VERSION : 0.1
// Die Funktion wird in einer Sprungleiste mit folgenden Schritten bearbeitet:
// 0: Warten, bis RT gedreht hat (nur danach ist Kettenentlastung notwendig)
// 1: Warten, bis BA Hand und keine Bewegung angefordert
// 2: Wartezeit vor Entlastung der Kette
//    -> Schritt 3, falls Wartezeit abgelaufen
//    -> Schritt 1, falls Automatik erneut angewählt oder Rundtisch dreht
// 3: Entlastung der Kette mit Zeitüberwachung
//    -> Schritt 1, falls während der Entlastung Bewegung angefordert wird
//    -> Schritt 0, falls während der Entlastung Automatik angewählt wird
// 4: Spannen der Kette mit Zeitüberwachung
   VAR_INPUT
      IN_P_Kette : Bool;   // Eingang von Druckschalter des Kettenspanners
      IN_Timer_Stg_Kette : Timer;   // Timer für die Störungsbildung der Spannung der Laufketten
      IN_Timer_Kettenspanner : Timer;   // Timer für den allgemeinen Ablauf des Kettenspanners
      IN_DW_Wartezeit : S5Time;   // Zeitwert für die Wartezeit nach Rundtisch im Handbetrieb
      IN_DW_Entlastungszeit : S5Time;   // Zeitwert für die Entlastungszeit der Kette
      IN_RT_dreht : Bool;   // Signal das sich der Rundtisch in Bewegung befindet
      IN_Steuerspannung : Bool;   // Signal Steuerspannung Eingeschaltet und Not- Aus entriegelt
      IN_Automatik_Stop_ok : Bool;   // Eingang das die Sicherheitseinrichtungen quittiert sind
      IN_Hydraulik_ok : Bool;   // Signal bei hydraulischen Kettenspannern das die Hydraulik bereit ist
      IN_Kettenspannung_noetig : Bool;   // Signal von extern das keine Kettenspannung nötig ist
      IN_Betriebsart_Automatik : Bool;   // Die Anlage befindet sich im Automatik- Betrieb
      IN_Start_Anlagenbetrieb : Bool;   // Die Anlage befindet sich in der Vorbereitung zum Produktionsbetrieb
      IN_Anlagenbetrieb : Bool;   // Die Anlage befindet sich im Produktionsbetrieb
      IN_Reset_fault_Fkt : Bool;   // Signal zum quittieren der Störungen innerhalb der einzelnen Funktionsbausteine
   END_VAR
   VAR_OUTPUT
      OUT_V_Entlastung : Bool;   // Ausgang für die Ansteuerung des Ketten- Entlastungs- Ventils
   END_VAR
   VAR_IN_OUT
      IO_Status : "UDT_RT_Kettenspanner";   // Speichern der Kettenentlastungs- Zustände für das Programm
   END_VAR
   VAR_TEMP
      Temp_IO_Status : "UDT_RT_Kettenspanner";   // Temporärer Kettenentlastungs- Status für die interne Bearbeitung des Bausteins
      ERROR_CODE : Int;   // Störungszustand der Systemfunktion "BLKMOV" Blockmove
      Anyzeiger : ANY;   // Zeiger zum Kopieren der Bereiche "IO_Status" und "Temp_IO_Status"
      Entlastung_starten : Bool;   // Zwischenmerker zum starten des Ablaufes der Kettenentspannung
   END_VAR
BEGIN

REGION Network 1: Gesicherte Daten einbinden
         LAR1;
         L;
         LAR2;
   //
         L     W#16#1002;  // Bytes
         T     W[AR1, P#0.0];
         L     2;  // Anzahl Bytes
         T     W[AR1, P#2.0];
         L     W[AR2, P#0.0];  // Baustein Nr.
         T     W[AR1, P#4.0];
         L     D[AR2, P#2.0];  // Datenanfang
         T     D[AR1, P#6.0];
   //
         CALL  BLKMOV
         ( SRCBLK  := #Anyzeiger,
           RET_VAL := #ERROR_CODE,
           DSTBLK  := #Temp_IO_Status
         );
   //
END_REGION

REGION Network 2: Stoerungen quittieren
         A     #IN_Reset_fault_Fkt;
         R     #Temp_IO_Status.STG_Entlastung;
         R     #Temp_IO_Status.STG_Druckaufbau;
END_REGION

REGION Network 3: Sprungleiste
         L     #Temp_IO_Status.Schrittnummer;
         JL    del;
         JU    dreh;  // 0: Warten, bis Rundtisch dreht
         JU    wrth;  // 1: Warten auf Betriebsart Hand + RT steht
         JU    wart;  // 2: Wartezeit vor Entlastung
         JU    entl;  // 3: Kettenentlastung
         JU    span;  // 4: Kette spannen
   del:  L     0;
         T     #Temp_IO_Status.Schrittnummer;
         CLR;
         =     #Temp_IO_Status.V_Entlastung;
         SP    #IN_Timer_Kettenspanner;
         SP    #IN_Timer_Stg_Kette;
         BEU;
END_REGION

REGION Network 4: 0: Warten, bis Rundtisch in Automatik gedreht hat
   dreh: ON    #IN_RT_dreht;
         ON    #IN_Anlagenbetrieb;
         JC    ende;
         L     1;
         T     #Temp_IO_Status.Schrittnummer;
         JU    ende;
END_REGION

REGION Network 5: 1: Warten, bis Automatik beendet und keine Bewegung läuft
   wrth: O     #IN_RT_dreht;
         O     #IN_Betriebsart_Automatik;
         JC    ende;
         L     2;
         T     #Temp_IO_Status.Schrittnummer;
         JU    ende;
END_REGION

REGION Network 6: 2: Wartezeit vor Kettenentlastung
   wart: SET;
         L     #IN_DW_Wartezeit;
         SD    #IN_Timer_Kettenspanner;
         L     1;
         O     #IN_RT_dreht;
         O     #IN_Start_Anlagenbetrieb;
         O     #IN_Anlagenbetrieb;
         JC    trnr;
         L     3;
         A     #IN_Timer_Kettenspanner;
         JC    trnr;
         JU    ende;
   trnr: T     #Temp_IO_Status.Schrittnummer;
         CLR;
         SP    #IN_Timer_Kettenspanner;
END_REGION

REGION Network 7: 3: Kettenentlastung
   entl: A     #IN_Steuerspannung;
         A     #IN_Automatik_Stop_ok;
         AN    #IN_RT_dreht;
         AN    #IN_Betriebsart_Automatik;
         AN    #IN_Kettenspannung_noetig;
         =     #Entlastung_starten;
         L     #IN_DW_Entlastungszeit;
         SP    #IN_Timer_Kettenspanner;
   //
         A     #Entlastung_starten;
         A     #IN_Timer_Kettenspanner;
         =     #Temp_IO_Status.V_Entlastung;
   //
         L     1;
         AN    #Entlastung_starten;
         JC    trn2;
         L     4;
         A     #Entlastung_starten;
         AN    #Temp_IO_Status.V_Entlastung;
         JC    trn2;
         JU    ende;
   trn2: T     #Temp_IO_Status.Schrittnummer;
         CLR;
         SP    #IN_Timer_Kettenspanner;
         JU    ende;
END_REGION

REGION Network 8: 4: Kette Spannen
   span: R     #Temp_IO_Status.V_Entlastung;
         L     0;
         T     #Temp_IO_Status.Schrittnummer;
END_REGION

REGION Network 9: Ende
   ende: A     #Temp_IO_Status.V_Entlastung;
         A     #IN_P_Kette;
         O;
         AN    #Temp_IO_Status.V_Entlastung;
         AN    #IN_P_Kette;
         A     #IN_Hydraulik_ok;
         L     S5T#10S;
         SD    #IN_Timer_Stg_Kette;
   //
         A     #IN_Timer_Stg_Kette;
         A     #Temp_IO_Status.V_Entlastung;
         S     #Temp_IO_Status.STG_Entlastung;
   //
         A     #IN_Timer_Stg_Kette;
         AN    #Temp_IO_Status.V_Entlastung;
         S     #Temp_IO_Status.STG_Druckaufbau;
   //
         AN    #Temp_IO_Status.V_Entlastung;
         A     #IN_P_Kette;
         =     #Temp_IO_Status.Kette_gespannt;
END_REGION

REGION Network 10: Ansteuerung des Entlanstungsventils
         A     #Temp_IO_Status.V_Entlastung;
         =     #OUT_V_Entlastung;
END_REGION

REGION Network 11: Daten sichern
         CALL  BLKMOV
         ( SRCBLK  := #Temp_IO_Status,
           RET_VAL := #ERROR_CODE,
           DSTBLK  := #Anyzeiger
         );
   //
END_REGION
END_FUNCTION

FUNCTION "FC1045_getStationRW" : Int   // FC1045, SCL
TITLE = Stationsnummer bestimmen
{ S7_Optimized_Access := 'FALSE' }
AUTHOR : AJ
VERSION : 2.0
// Stationsnummer bestimmen,anhand des Positionsistwert
// KNOW_HOW_PROTECT
   VAR_INPUT
      Anzahl_Segmente : Int;   // Wieviel Segmente hat der RT?
      Maxwert : DInt;   // Eine Umdrehung hat soviele Grad oder Inc (360°)
      Offset : DInt;   // Verschiebung um soviel Grad
      Istwert : DInt;   // Vom Umrichter
      SegmenteReverse : Bool;   // Haben Segmente absteigende Reihenfolge? (10,9,8,...)
   END_VAR
   VAR_TEMP
      anfang : Int;
      ende : Int;
      schrittweite : Int;
      laufvariable : Int;
      Segmentgroesse : DInt;
      Vergleichswert1 : DInt;
      Vergleichswert2 : DInt;
      IstwertPlus : DInt;
      Offset_temp : DInt;
      result : Int;
   END_VAR
BEGIN



                     #anfang:= 1;
                     #schrittweite:=1; 
                     #ende:= #Anzahl_Segmente;
                     #laufvariable:=1;

                     #Segmentgroesse:= #Maxwert/#Anzahl_Segmente;
              // Offset begrenzen auf Segmentbreite
                     IF  #Offset < (#Segmentgroesse-20)  THEN
                     #Offset_temp:=#Offset;
                     ELSE
                     #Offset_temp:=#Segmentgroesse-20;
                     END_IF;
               // Istwert mit Offset verrechnen
                     #IstwertPlus:=#Istwert+#Offset_temp;
                       IF  #IstwertPlus < 3600 THEN
                       #IstwertPlus:= #IstwertPlus;
                       ELSE
                       #IstwertPlus:= #IstwertPlus-#Maxwert;                    
                       END_IF;  



                     FOR #laufvariable := #anfang TO #ende BY #schrittweite DO
                          #Vergleichswert1:= (#laufvariable-1)*#Segmentgroesse;
                          #Vergleichswert2:= #laufvariable*#Segmentgroesse;


                           IF  #IstwertPlus >= #Vergleichswert1 AND #IstwertPlus < #Vergleichswert2   THEN

                               IF #SegmenteReverse = false THEN
                               #result:=#laufvariable;
                               ELSE
                               #result:=#Anzahl_Segmente+1-#laufvariable;
                               END_IF;


                           EXIT;


                            END_IF;

                      END_FOR;

   #FC1045_getStationRW:= #result;
END_FUNCTION

FUNCTION "FC1046_SegmInStation" : Void   // FC1046, SCL
{ S7_Optimized_Access := 'FALSE' }
VERSION : 0.1
   VAR_INPUT
      IN_Amount_Segment : Int;
   END_VAR
   VAR_TEMP
      N : Int;   // Laufvariable
      Z : Int;
   END_VAR
BEGIN
   // Schieben der einzelnen Segmentnummern in die Sationen
   // Aktuell nur in Uhrzeigersinn und in aufsteigender Reihenfolge

   IF "DB1001_TT_State".SegmentInfo[1].SegmentNo <> "DB1001_TT_State".Segmentkennung.Seg_No_Stat_1 THEN

       "DB1001_TT_State".SegmentInfo[1].SegmentNo := "DB1001_TT_State".Segmentkennung.Seg_No_Stat_1;
       #Z := "DB1001_TT_State".SegmentInfo[1].SegmentNo;

       FOR #N := 2 TO #IN_Amount_Segment DO
           IF #Z > 1 THEN
               "DB1001_TT_State".SegmentInfo[#N].SegmentNo := #Z - 1;
           ELSE
               "DB1001_TT_State".SegmentInfo[#N].SegmentNo := #Z + #IN_Amount_Segment - 1;
           END_IF;
           #Z := #Z - 1;
       END_FOR;


   //    // Zählt falsch herum!!
       //    "DB1001_RT".SegmentNoinStation[1] := "DB1001_RT".Segmentkennung.Seg_No_Stat_1;
       //    #Z := "DB1001_RT".SegmentNoinStation[1];

       //    FOR #N := 2 TO #IN_Amount_Segment DO
       //       IF #Z < #IN_Amount_Segment THEN
       //         "DB1001_RT".SegmentNoinStation[#N] := #Z + 1;
       //    ELSE
       //        "DB1001_RT".SegmentNoinStation[#N] := #Z - #IN_Amount_Segment + 1;
       //    END_IF;
       //    #Z := #Z + 1;
       //END_FOR;

   END_IF;

   FOR #N := 1 TO #IN_Amount_Segment DO
       IF "DB1001_TT_State".SegmentInfo[#N].SegmentNo > 0 THEN
           "DB1001_TT_State".SegmentInfo[#N].Enable := "DB1051_TT_SegValue".Station["DB1001_TT_State".SegmentInfo[#N].SegmentNo].FoamingEnable;
           "DB1001_TT_State".SegmentInfo[#N].ShotDone := "DB1001_TT_State".SegmentWithFoam["DB1001_TT_State".SegmentInfo[#N].SegmentNo];
           "DB1001_TT_State".SegmentInfo[#N].FoamingProgram := "DB1051_TT_SegValue".Station["DB1001_TT_State".SegmentInfo[#N].SegmentNo].FoamingProg;
           "DB1001_TT_State".SegmentInfo[#N].Status := "DB1001_TT_State".SegmentStatus["DB1001_TT_State".SegmentInfo[#N].SegmentNo];
       ELSE
           "DB1001_TT_State".SegmentInfo[#N].Enable := 0;
           "DB1001_TT_State".SegmentInfo[#N].ShotDone := 0;
           "DB1001_TT_State".SegmentInfo[#N].FoamingProgram := 0;
           "DB1001_TT_State".SegmentInfo[#N].Status := 0;
       END_IF;
   END_FOR;
END_FUNCTION

FUNCTION "FC1051_TT_Segment" : Void   // FC1051, STL
{ S7_Optimized_Access := 'TRUE' }
VERSION : 0.1
BEGIN

REGION Network 1: No Foaming
         A     "DB1001_TT_State".IPOS.Status.RT_in_Position;
         A     "Button_without_foam";
         S     "DB1001_TT_State".Bits.NoFoamingButton;

         AN    "DB1001_TT_State".IPOS.Status.RT_in_Position;
         R     "DB1001_TT_State".Bits.NoFoamingButton;

   //      U     "DB1001_TT_State".Bits.NoFoamingButton
   //      =     "TT_H_WithoutFoam"
END_REGION

REGION Network 2: Emptying
         A     "Button_TT_empty";
         S     "DB1001_TT_State".Bits.TTEmptying;

         AN    "DB1001_TT_State".BA_Anlage.Produktion;
         R     "DB1001_TT_State".Bits.TTEmptying;

         AN    "DB1001_TT_State".SegmentWithFoam[1];
         AN    "DB1001_TT_State".SegmentWithFoam[2];
         AN    "DB1001_TT_State".SegmentWithFoam[3];
         AN    "DB1001_TT_State".SegmentWithFoam[4];
         AN    "DB1001_TT_State".SegmentWithFoam[5];
         AN    "DB1001_TT_State".SegmentWithFoam[6];
         AN    "DB1001_TT_State".SegmentWithFoam[7];
         AN    "DB1001_TT_State".SegmentWithFoam[8];
         A     "DB1001_TT_State".Bits.TTEmptying;
         =     "DB1001_TT_State".Bits.StopAfterEmpty;

         A     "DB1001_TT_State".Bits.TTEmptying;
         =     "LED_TT_empty";
END_REGION

REGION Network 3: Interface TT <-> RS
   //-----
         O     "DB005_RS<->Extern".MC_Interface[1].Data_to_MC.Shot_end;
         =     "DB1001_TT_State".SegmentShotEnds[1];
         =     "DB1001_TT_State".SegmentShotEnds[2];
         =     "DB1001_TT_State".SegmentShotEnds[3];
         =     "DB1001_TT_State".SegmentShotEnds[4];
         =     "DB1001_TT_State".SegmentShotEnds[5];
         =     "DB1001_TT_State".SegmentShotEnds[6];
         =     "DB1001_TT_State".SegmentShotEnds[7];
         =     "DB1001_TT_State".SegmentShotEnds[8];
   //-----
         O     "DB1001_TT_State".SegmentPreperationFoaming[1];
         O     "DB1001_TT_State".SegmentPreperationFoaming[2];
         O     "DB1001_TT_State".SegmentPreperationFoaming[3];
         O     "DB1001_TT_State".SegmentPreperationFoaming[4];
         O     "DB1001_TT_State".SegmentPreperationFoaming[5];
         O     "DB1001_TT_State".SegmentPreperationFoaming[6];
         O     "DB1001_TT_State".SegmentPreperationFoaming[7];
         O     "DB1001_TT_State".SegmentPreperationFoaming[8];
         =     "DB005_RS<->Extern".MC_Interface[1].Data_from_MC.Shot_preperation;
   //-----
         O     "DB1001_TT_State".SegmentEnableFoaming[1];
         O     "DB1001_TT_State".SegmentEnableFoaming[2];
         O     "DB1001_TT_State".SegmentEnableFoaming[3];
         O     "DB1001_TT_State".SegmentEnableFoaming[4];
         O     "DB1001_TT_State".SegmentEnableFoaming[5];
         O     "DB1001_TT_State".SegmentEnableFoaming[6];
         O     "DB1001_TT_State".SegmentEnableFoaming[7];
         O     "DB1001_TT_State".SegmentEnableFoaming[8];
         =     "DB005_RS<->Extern".MC_Interface[1].Data_from_MC.Shot_release;
   //-----
END_REGION
END_FUNCTION

FUNCTION "FC1156_FlowPressMH_Instance" : Void   // FC1156, SCL
{ S7_Optimized_Access := 'FALSE' }
VERSION : 0.1
   VAR_INPUT
      IN_MachineNo : Int;
      IN_MixingHeadNo : Int;
      IN_AmountMHConnections : Byte;
      IN_Cycle : Bool;
      IN_ReducedRecirculation : Bool;
      IN_LPRecirculation : Bool;
      IN_HPRecirculation : Bool;
      IN_PauseTime : Bool;
      IN_Reset_Fault : Bool;
   END_VAR
   VAR_IN_OUT
      IO_FaultWrongAssignment : Bool;   // Wrong assignment of tank to pump or pump to mixinghead
      IO_Fault_Level_1 : Bool;
      IO_New_Fault : Bool;
   END_VAR
   VAR_TEMP
      Tmp_ComponentNo : Int;
      TmpPressure : Word;
      TmpPumpNo : Int;
      TmpFlow : DInt;
      TmpShotActive : Bool;
      TmpFlowQPB : DInt;
      Tmp_ShotConn : Word;
      Tmp_ShotComp : Word;
      Tmp_CompNoShot : Word;
      Tmp_ShotCompShift : Word;
      Tmp_AmountMHConnections : Int;
      i : Int;
      Test : Int;
      Test2 : Int;
   END_VAR
BEGIN
   // Initialization temporary variables
   #Tmp_ShotConn := 0;
   #Tmp_ShotComp := 0;
   #TmpShotActive := FALSE;
   #Tmp_AmountMHConnections := #IN_AmountMHConnections;  // This should be a input parameter

   // Reset Fault
   IF #IN_Reset_Fault THEN
      #IO_FaultWrongAssignment := FALSE;
   END_IF;

   // For loop over all mixinghead connections
   FOR #i := 1 TO #Tmp_AmountMHConnections DO

       // Get pump no. connected with mixinghead connector
       #TmpPumpNo       := "DB704_MH_Value".Mixinghead[#IN_MixingHeadNo].MH_Connection[#i].Pump_No;
       #Tmp_ComponentNo := "DB753_MeteringPump".Pump[#TmpPumpNo].TankNo;

       // Wrong assignment of tank to pump or pump to mixinghead
       IF #TmpPumpNo = 0 OR #Tmp_ComponentNo = 0  AND NOT #IO_FaultWrongAssignment THEN
         #IO_FaultWrongAssignment := TRUE;
         #IO_Fault_Level_1        := TRUE;
         #IO_New_Fault            := TRUE;
         EXIT;
       END_IF;

       // If at the pump no 2- Point- Adjustment seleced delet the MH values
       IF "DB753_MeteringPump".Pump[#TmpPumpNo].With_2Point = 0 THEN
         "DB704_MH_Value".Mixinghead[#IN_MixingHeadNo].MH_Connection[#i].Red_2Point_Flow := 0;
         "DB704_MH_Value".Mixinghead[#IN_MixingHeadNo].MH_Connection[#i].LP_2Point_Flow := 0;
         "DB704_MH_Value".Mixinghead[#IN_MixingHeadNo].MH_Connection[#i].HP_2Point_Flow := 0;
       END_IF;

       // Get flow values at reduced, low pressure and high pressure cycle
       IF #IN_ReducedRecirculation AND NOT #IN_PauseTime THEN
         "DB613_Komponent_State".FlowPump[#TmpPumpNo] := "DB704_MH_Value".Mixinghead[#IN_MixingHeadNo].MH_Connection[#i].Flow_red_Circ;
         //"DB613_Komponent_State".MeteringPump[#TmpPumpNo]."2PointAdjustmentSelected" := "DB704_MH_Value".Mixinghead[#IN_MixingHeadNo].MH_Connection[#i].Red_2Point_Flow;
       ELSIF #IN_LPRecirculation AND NOT #IN_PauseTime THEN
         "DB613_Komponent_State".FlowPump[#TmpPumpNo] := "DB704_MH_Value".Mixinghead[#IN_MixingHeadNo].MH_Connection[#i].Flow_LP_Circ;
         //"DB613_Komponent_State".MeteringPump[#TmpPumpNo]."2PointAdjustmentSelected" := "DB704_MH_Value".Mixinghead[#IN_MixingHeadNo].MH_Connection[#i].LP_2Point_Flow;
       ELSIF #IN_HPRecirculation THEN
         "DB613_Komponent_State".FlowPump[#TmpPumpNo] := "DB704_MH_Value".Mixinghead[#IN_MixingHeadNo].MH_Connection[#i].Flow_HP_Circ; 
         //"DB613_Komponent_State".MeteringPump[#TmpPumpNo]."2PointAdjustmentSelected" := "DB704_MH_Value".Mixinghead[#IN_MixingHeadNo].MH_Connection[#i].HP_2Point_Flow;
       ELSE
         "DB613_Komponent_State".FlowPump[#TmpPumpNo] := 0;
         //"DB613_Komponent_State".MeteringPump[#TmpPumpNo]."2PointAdjustmentSelected" := 0;
       END_IF;

       // IS get flow of pump at cycle and set component active 
       IF #TmpPumpNo > 0 AND #IN_Cycle THEN
           IF "DB619_State_MPart".ShotMa[#IN_MachineNo].ShotData.Flow[#i] > 0 THEN
           #TmpShotActive := TRUE;
           // Pressure and flow at connection 1 mixinghead at foaming cycle
           "DB613_Komponent_State".FlowPump[#TmpPumpNo]  := "DB619_State_MPart".ShotMa[#IN_MachineNo].ShotData.Flow[#i];
           "DB604_PV_Mixinghead".Mixinghead[#IN_MixingHeadNo].Pressure_Connection[#i].PV_SetV.Value  := "DB619_State_MPart".ShotMa[#IN_MachineNo].ShotData.Pressure[#i];
           //"DB613_Komponent_State".MeteringPump[#TmpPumpNo]."2PointAdjustmentSelected" := "DB619_State_MPart".ShotMa[#IN_MachineNo].ShotData."2PointAdjustment"[#i];
         ELSE
           // If Flow = 0 take the high pressure flow
           "DB613_Komponent_State".FlowPump[#TmpPumpNo] := "DB704_MH_Value".Mixinghead[#IN_MixingHeadNo].MH_Connection[#i].Flow_HP_Circ; 
           //"DB613_Komponent_State".MeteringPump[#TmpPumpNo]."2PointAdjustmentSelected" := "DB704_MH_Value".Mixinghead[#IN_MixingHeadNo].MH_Connection[#i].HP_2Point_Flow;
           #TmpShotActive := FALSE;
         END_IF;
       ELSE
         #TmpShotActive := FALSE;
       END_IF;



       // Set value for the flow controls
       "DB608_PV_Metering".Metering[#TmpPumpNo].Flow.PV_SetV.Value := "DB613_Komponent_State".FlowPump[#TmpPumpNo];

       // Get flow and pressure for quick pressure build up
       IF #IN_Cycle  OR #IN_HPRecirculation THEN
         "DB613_Komponent_State".FlowPumpQPB[#TmpPumpNo]      := "DB704_MH_Value".Mixinghead[#IN_MixingHeadNo].MH_Connection[#i].FlowQPB;
         "DB613_Komponent_State".PressurePumpQPB[#TmpPumpNo]  := "DB704_MH_Value".Mixinghead[#IN_MixingHeadNo].MH_Connection[#i].PressureQPB;
       ELSE
         "DB613_Komponent_State".FlowPumpQPB[#TmpPumpNo]      := "DB704_MH_Value".Mixinghead[#IN_MixingHeadNo].MH_Connection[#i].FlowQPB;; // 0;
         "DB613_Komponent_State".PressurePumpQPB[#TmpPumpNo]  := "DB704_MH_Value".Mixinghead[#IN_MixingHeadNo].MH_Connection[#i].PressureQPB; // 0;
       END_IF;

       // Set component bit if used at this shot and connection bit used at this shot
       IF #TmpShotActive  THEN
         #Tmp_CompNoShot    := 1;
         #Tmp_ShotCompShift := SHL(IN :=#Tmp_CompNoShot, N := #TmpPumpNo -1);
         #Tmp_ShotComp      := #Tmp_ShotComp OR #Tmp_ShotCompShift;

         #Tmp_ShotConn := #Tmp_ShotConn OR #Tmp_ShotComp;// INT_TO_WORD(#i); // Connection number
       END_IF;

   END_FOR;


   // SetValue for the mixinghead ratio
   // 
   // SetValue for the mixinghead ratio

   IF "DB613_Komponent_State".MeteringPump[1].Metering_to_PUC = TRUE AND "DB614_MH_State".MH_Status[1].Switch_Testshot_B_ON_OFF = FALSE AND "DB608_PV_Metering".Metering[1].Flow.PV_ActV.Value > 0 THEN
       "DB608_PV_Metering".Metering[1].MixingRatio.PV_ActV.Value :=
       "DB608_PV_Metering".Metering[1].Flow.PV_ActV.Value * REAL#100.0 /
       "DB608_PV_Metering".Metering[1].Flow.PV_ActV.Value;
   ELSE
       "DB608_PV_Metering".Metering[1].MixingRatio.PV_ActV.Value := 100.0;
   END_IF;

   IF "DB614_MH_State".MH_Status[1].Switch_Testshot_B_ON_OFF = TRUE THEN

       "DB608_PV_Metering".Metering[1].MixingRatio.PV_ActV.Value := 0.0;

   END_IF;

   IF "DB613_Komponent_State".MeteringPump[2].Metering_to_PUC = TRUE AND "DB614_MH_State".MH_Status[1].Switch_Testshot_A_ON_OFF = FALSE AND "DB608_PV_Metering".Metering[2].Flow.PV_ActV.Value > 0 THEN
       "DB608_PV_Metering".Metering[2].MixingRatio.PV_ActV.Value :=
       "DB608_PV_Metering".Metering[2].Flow.PV_ActV.Value * REAL#100.0 /
       "DB608_PV_Metering".Metering[1].Flow.PV_ActV.Value;
   ELSE
       "DB608_PV_Metering".Metering[2].MixingRatio.PV_ActV.Value := 100.0;
   END_IF;

   IF "DB614_MH_State".MH_Status[1].Switch_Testshot_A_ON_OFF = TRUE THEN

       "DB608_PV_Metering".Metering[2].MixingRatio.PV_ActV.Value := 0.0;

   END_IF;

   "DB608_PV_Metering".Metering[3].MixingRatio.PV_ActV.Value :=
   "DB608_PV_Metering".Metering[3].Flow.PV_ActV.Value * REAL#100.0 /
   "DB608_PV_Metering".Metering[1].Flow.PV_ActV.Value;

   "DB608_PV_Metering".Metering[4].MixingRatio.PV_ActV.Value :=
   "DB608_PV_Metering".Metering[4].Flow.PV_ActV.Value * REAL#100.0 /
   "DB608_PV_Metering".Metering[1].Flow.PV_ActV.Value;

   "DB608_PV_Metering".Metering[5].MixingRatio.PV_ActV.Value :=
   "DB608_PV_Metering".Metering[5].Flow.PV_ActV.Value * REAL#100.0 /
   "DB608_PV_Metering".Metering[1].Flow.PV_ActV.Value;

   "DB608_PV_Metering".Metering[6].MixingRatio.PV_ActV.Value :=
   "DB608_PV_Metering".Metering[6].Flow.PV_ActV.Value * REAL#100.0 /
   "DB608_PV_Metering".Metering[1].Flow.PV_ActV.Value;

   "DB608_PV_Metering".Metering[7].MixingRatio.PV_ActV.Value :=
   "DB608_PV_Metering".Metering[7].Flow.PV_ActV.Value * REAL#100.0 /
   "DB608_PV_Metering".Metering[1].Flow.PV_ActV.Value;

   "DB608_PV_Metering".Metering[8].MixingRatio.PV_ActV.Value :=
   "DB608_PV_Metering".Metering[8].Flow.PV_ActV.Value * REAL#100.0 /
   "DB608_PV_Metering".Metering[1].Flow.PV_ActV.Value;

   "DB608_PV_Metering".Metering[9].MixingRatio.PV_ActV.Value :=
   "DB608_PV_Metering".Metering[9].Flow.PV_ActV.Value * REAL#100.0 /
   "DB608_PV_Metering".Metering[1].Flow.PV_ActV.Value;

   "DB608_PV_Metering".Metering[10].MixingRatio.PV_ActV.Value :=
   "DB608_PV_Metering".Metering[10].Flow.PV_ActV.Value * REAL#100.0 /
   "DB608_PV_Metering".Metering[1].Flow.PV_ActV.Value;

   "DB608_PV_Metering".Metering[11].MixingRatio.PV_ActV.Value :=
   "DB608_PV_Metering".Metering[11].Flow.PV_ActV.Value * REAL#100.0 /
   "DB608_PV_Metering".Metering[1].Flow.PV_ActV.Value;

   "DB608_PV_Metering".Metering[12].MixingRatio.PV_ActV.Value :=
   "DB608_PV_Metering".Metering[12].Flow.PV_ActV.Value * REAL#100.0 /
   "DB608_PV_Metering".Metering[1].Flow.PV_ActV.Value;


   "DB619_State_MPart".ShotMa[#IN_MachineNo].ShotData.Comp_at_Shot := #Tmp_ShotConn;
END_FUNCTION

FUNCTION "FC1500_ShotDataToMC" : Void   // FC1500, STL
TITLE = Shot data to MCs
{ S7_Optimized_Access := 'FALSE' }
VERSION : 0.1
   VAR_TEMP
      RetVal : Int;
      nullbyte : Byte;
      RetValSFC : Int;
   END_VAR
BEGIN

REGION Network 1: Read data from bus
   // MC1
   //      CALL  DPRD_DAT
   //         LADDR   :="PN-PN-Coupler_PU_MC1~IN___2_Byte"
   //         RET_VAL :=#RetValSFC
   //         RECORD  :="DB1500_ShotDataToMC".ShotData_MC[1].Data_from_MC
   // MC2
   //      CALL  DPRD_DAT
   //         LADDR   :="PN-PN-Coupler_PU_MC2~IN___2_Byte"
   //         RET_VAL :=#RetValSFC
   //         RECORD  :="DB1500_ShotDataToMC".ShotData_MC[2].Data_from_MC
   // MC3
   // CALL  DPRD_DAT
   //         LADDR   :="PN-PN-Coupler_MC3~IN___2_Byte"
   //         RET_VAL :=#RetValSFC
   //         RECORD  :="DB1500_ShotDataToMC".ShotData_MC[3].Data_from_MC
   // MC4
   // CALL  DPRD_DAT
   //         LADDR   :="PN-PN-Coupler_MC4~IN___2_Byte"
   //         RET_VAL :=#RetValSFC
   //         RECORD  :="DB1500_ShotDataToMC".ShotData_MC[4].Data_from_MC
END_REGION

REGION Network 2: Communication control
   // If the mouldcarrier doesn't read its shotdata after two seconds it will reset 
   // automatically
   // Handshake with the mouldcarrier 01
         AN    "DB1500_ShotDataToMC".ShotData_MC[1].Data_from_MC.Communication.Data_read;
         A     "DB1500_ShotDataToMC".ShotData_MC[1].Data_to_MC.Communication.New_Data;
         L     S5T#2S;
         SD    "TM_FLT_Com_DataShot_MC01";

         O     "DB1500_ShotDataToMC".ShotData_MC[1].Data_from_MC.Communication.Data_read;
         O     "TM_FLT_Com_DataShot_MC01";
         R     "DB1500_ShotDataToMC".ShotData_MC[1].Data_from_MC.Communication.Data_read;
         R     "DB1500_ShotDataToMC".ShotData_MC[1].Data_to_MC.Communication.New_Data;
         R     "TM_FLT_Com_DataShot_MC01";

   // Handshake with the mouldcarrier 02
         AN    "DB1500_ShotDataToMC".ShotData_MC[2].Data_from_MC.Communication.Data_read;
         A     "DB1500_ShotDataToMC".ShotData_MC[2].Data_to_MC.Communication.New_Data;
         L     S5T#2S;
         SD    "TM_FLT_Com_DataShot_MC02";

         O     "DB1500_ShotDataToMC".ShotData_MC[2].Data_from_MC.Communication.Data_read;
         O     "TM_FLT_Com_DataShot_MC02";
         R     "DB1500_ShotDataToMC".ShotData_MC[2].Data_from_MC.Communication.Data_read;
         R     "DB1500_ShotDataToMC".ShotData_MC[2].Data_to_MC.Communication.New_Data;
         R     "TM_FLT_Com_DataShot_MC02";

   // Handshake with the mouldcarrier 03
         AN    "DB1500_ShotDataToMC".ShotData_MC[3].Data_from_MC.Communication.Data_read;
         A     "DB1500_ShotDataToMC".ShotData_MC[3].Data_to_MC.Communication.New_Data;
         L     S5T#2S;
         SD    "TM_FLT_Com_DataShot_MC03";

         O     "DB1500_ShotDataToMC".ShotData_MC[3].Data_from_MC.Communication.Data_read;
         O     "TM_FLT_Com_DataShot_MC03";
         R     "DB1500_ShotDataToMC".ShotData_MC[3].Data_from_MC.Communication.Data_read;
         R     "DB1500_ShotDataToMC".ShotData_MC[3].Data_to_MC.Communication.New_Data;
         R     "TM_FLT_Com_DataShot_MC03";

   // Handshake with the mouldcarrier 04
         AN    "DB1500_ShotDataToMC".ShotData_MC[4].Data_from_MC.Communication.Data_read;
         A     "DB1500_ShotDataToMC".ShotData_MC[4].Data_to_MC.Communication.New_Data;
         L     S5T#2S;
         SD    "TM_FLT_Com_DataShot_MC04";  // ""

         O     "DB1500_ShotDataToMC".ShotData_MC[4].Data_from_MC.Communication.Data_read;
         O     "TM_FLT_Com_DataShot_MC04";
         R     "DB1500_ShotDataToMC".ShotData_MC[4].Data_from_MC.Communication.Data_read;
         R     "DB1500_ShotDataToMC".ShotData_MC[4].Data_to_MC.Communication.New_Data;
         R     "TM_FLT_Com_DataShot_MC04";
END_REGION

REGION Network 3: Shot start --> the set values will be transfer to the interface
         A     "DB619_State_MPart".Cycle[1].ShotRuns;
         FP    "HF_new_setvalue_Of_ShotData";
         A     "DB123_MH_IO_Signals".MH[1].IN.MH_Auto_Mode;
         JCN   newSetData;

   newSetData:NOP   0;
END_REGION

REGION Network 4: Shot finished --> the atual values will be transfer to the interface
         A     "M_NewShotDataToMC";
         FP    "HF_new_shot_data";
         JCN   newData;
END_REGION

REGION Network 5: Shot data to buffer
   //----------------------------------------------------------------
   // Actual station number
   //----------------------------------------------------------------
         L     "DB919_ShotResultMach".ShotResult_Ma[1].General.StationNo;
         T     "DB1500_ShotDataToMC".ShotData_MC[0].Data_to_MC.Shot_data.Station_No;
   //----------------------------------------------------------------
   // Actual mixing head number
   //----------------------------------------------------------------
         L     "DB919_ShotResultMach".ShotResult_Ma[1].General.MH_No;
         T     "DB1500_ShotDataToMC".ShotData_MC[0].Data_to_MC.Shot_data.MH_No;
   //----------------------------------------------------------------
   // Actual shot no
   //----------------------------------------------------------------
         L     "DB919_ShotResultMach".ShotResult_Ma[1].General.PartID;
         T     "DB1500_ShotDataToMC".ShotData_MC[0].Data_to_MC.Shot_data.Shot_No;
   //----------------------------------------------------------------
   // Date and Time Shot end
   //----------------------------------------------------------------
         CALL  MOVE
         ( IN  := "DB919_ShotResultMach".ShotResult_Ma[1].General.DateTime,
           OUT := "DB1500_ShotDataToMC".ShotData_MC[0].Data_to_MC.Shot_data.DateTime
         );

   //----------------------------------------------------------------
   // values of the shot time
   //----------------------------------------------------------------
   // actual value [1/1 ms]
         L     "DB919_ShotResultMach".ShotResult_Ma[1].General.FoamingTime;
         T     "DB1500_ShotDataToMC".ShotData_MC[0].Data_to_MC.Shot_data.ShotTime_act;

   // set value [1/1 ms]
         L     "DB619_State_MPart".ShotMa[1].Tool.Shot[1].FoamingTime;
         T     "DB1500_ShotDataToMC".ShotData_MC[0].Data_to_MC.Shot_data.ShotTime_set;
   //----------------------------------------------------------------
   // values mixinghead shot weight
   //----------------------------------------------------------------
   // ActValue totally [1/1 g]
         L     "DB919_ShotResultMach".ShotResult_Ma[1].General.PartWeight;
         T     "DB1500_ShotDataToMC".ShotData_MC[0].Data_to_MC.Shot_data.ShotWeight_act;

   // SetValue totally [1/1 g]
         L     "DB619_State_MPart".ShotMa[1].Tool.Shot[1].PartWeight;
         T     "DB1500_ShotDataToMC".ShotData_MC[0].Data_to_MC.Shot_data.ShotWeight_set;
   //----------------------------------------------------------------
   // Actual values Mixinghead pressure component 01
   //----------------------------------------------------------------
   // actual value [1/1 bar]
         L     "DB919_ShotResultMach".ShotResult_Ma[1].Component.Comp[1].PressureMH;
         T     "DB1500_ShotDataToMC".ShotData_MC[0].Data_to_MC.Shot_data.Comp_act[1].Pressure_MH;

   // set value [1/1 bar]
         L     "DB619_State_MPart".ShotMa[1].Tool.Shot[1].Pressure[1];
         T     "DB1500_ShotDataToMC".ShotData_MC[0].Data_to_MC.Shot_data.Comp_set[1].Pressure_MH;

   //----------------------------------------------------------------
   // Actual values Mixinghead pressure component 02
   //----------------------------------------------------------------
   // actual value [1/10 bar]
         L     "DB919_ShotResultMach".ShotResult_Ma[1].Component.Comp[2].PressureMH;
         T     "DB1500_ShotDataToMC".ShotData_MC[0].Data_to_MC.Shot_data.Comp_act[2].Pressure_MH;

   // set value [1/1 bar]
         L     "DB619_State_MPart".ShotMa[1].Tool.Shot[1].Pressure[2];
         T     "DB1500_ShotDataToMC".ShotData_MC[0].Data_to_MC.Shot_data.Comp_set[2].Pressure_MH;

   //----------------------------------------------------------------
   // Actual values mixinghead temperature component C1
   //----------------------------------------------------------------
   // actual value [1/1 °C]
         L     "DB919_ShotResultMach".ShotResult_Ma[1].Component.Comp[1].TemperatureMH;
         T     "DB1500_ShotDataToMC".ShotData_MC[0].Data_to_MC.Shot_data.Comp_act[1].Temperature_MH;

   // set value[1/1°C]
         L     "DB604_PV_Mixinghead".Mixinghead[1].Temperature_Connection[1].PV_SetV.Value;
         T     "DB1500_ShotDataToMC".ShotData_MC[0].Data_to_MC.Shot_data.Comp_set[1].Temperature_MH;
   //----------------------------------------------------------------
   // Actual values mixinghead temperature component C2
   //----------------------------------------------------------------
   // actual value [1/1 °C]
         L     "DB919_ShotResultMach".ShotResult_Ma[1].Component.Comp[2].TemperatureMH;
         T     "DB1500_ShotDataToMC".ShotData_MC[0].Data_to_MC.Shot_data.Comp_act[2].Temperature_MH;

   // set value[1/1°C]
         L     "DB604_PV_Mixinghead".Mixinghead[1].Temperature_Connection[2].PV_SetV.Value;
         T     "DB1500_ShotDataToMC".ShotData_MC[0].Data_to_MC.Shot_data.Comp_set[2].Temperature_MH;
   //----------------------------------------------------------------
   // Actual values mixinghead flow component C1
   //----------------------------------------------------------------
   // actual value [1/1 g/s]
         L     "DB919_ShotResultMach".ShotResult_Ma[1].Component.Comp[1].Flow;
         T     "DB1500_ShotDataToMC".ShotData_MC[0].Data_to_MC.Shot_data.Comp_act[1].Flow;

   // set value [1/1 g/s]
         L     "DB619_State_MPart".ShotMa[1].ShotData.Flow[1];
         T     "DB1500_ShotDataToMC".ShotData_MC[0].Data_to_MC.Shot_data.Comp_set[1].Flow;
   //----------------------------------------------------------------
   // Actual values mixinghead flow component C2
   //----------------------------------------------------------------
   // actual value [1/1 g/s]
         L     "DB919_ShotResultMach".ShotResult_Ma[1].Component.Comp[2].Flow;
         T     "DB1500_ShotDataToMC".ShotData_MC[0].Data_to_MC.Shot_data.Comp_act[2].Flow;

   // setvalue [1/1 g/s]
         L     "DB619_State_MPart".ShotMa[1].ShotData.Flow[2];
         T     "DB1500_ShotDataToMC".ShotData_MC[0].Data_to_MC.Shot_data.Comp_set[2].Flow;


   // Set data valid
         SET;
         S     "HT_new_shot_data_valid";
         R     "M_NewShotDataToMC";

   newData:NOP   0;
END_REGION

REGION Network 6: Create jump order
   //----------------------------------
   // Prepare to send data MC 1
         A     "DB110_Interf_Program_M1".Status_IF[1].IF_is_on_1_Position;
         A     "DB619_State_MPart".Cycle[1].ShotRuns;
         FP    "M_FP_NewShotDataToMC_01";
   //      U     "DB123_MH_IO_Signals".MH[1].IN.MH_Auto_Mode
         S     "M_NewShotDataToMC_01";

         A     "M_NewShotDataToMC_01";
         A     "HT_new_shot_data_valid";
         AN    "M_WriteShotDataMC_01";
         S     "M_WriteShotDataMC_01";

   // Prepare to send data MC 2
         A     "DB110_Interf_Program_M1".Status_IF[2].IF_is_on_1_Position;
         A     "DB619_State_MPart".Cycle[1].ShotRuns;
         FP    "M_FP_NewShotDataToMC_02";
         A     "DB123_MH_IO_Signals".MH[1].IN.MH_Auto_Mode;
         S     "M_NewShotDataToMC_02";

         A     "M_NewShotDataToMC_02";
         A     "HT_new_shot_data_valid";
         AN    "M_WriteShotDataMC_02";
         S     "M_WriteShotDataMC_02";

   // Prepare to send data MC 3
         A     "DB110_Interf_Program_M1".Status_IF[3].IF_is_on_1_Position;
         A     "DB619_State_MPart".Cycle[1].ShotRuns;
         FP    "M_FP_NewShotDataToMC_03";
         A     "DB123_MH_IO_Signals".MH[1].IN.MH_Auto_Mode;
         S     "M_NewShotDataToMC_03";

         A     "M_NewShotDataToMC_03";
         A     "HT_new_shot_data_valid";
         AN    "M_WriteShotDataMC_03";
         S     "M_WriteShotDataMC_03";

   // Prepare to send data MC 4
         A     "DB110_Interf_Program_M1".Status_IF[4].IF_is_on_1_Position;
         A     "DB619_State_MPart".Cycle[1].ShotRuns;
         FP    "M_FP_NewShotDataToMC_04";
         A     "DB123_MH_IO_Signals".MH[1].IN.MH_Auto_Mode;
         S     "M_NewShotDataToMC_04";

         A     "M_NewShotDataToMC_04";
         A     "HT_new_shot_data_valid";
         AN    "M_WriteShotDataMC_04";
         S     "M_WriteShotDataMC_04";

   // If Interface 05 at the first postion (Testshot) reset the reminder "HT_new_shot_data_valid"
         A     "DB110_Interf_Program_M1".Status_IF[5].IF_is_on_1_Position;
         A     "DB619_State_MPart".Cycle[1].ShotRuns;
         FP    "M_FP_NewShotDataTestShot";
         A     "DB123_MH_IO_Signals".MH[1].IN.MH_Auto_Mode;
         S     "M_NewShotDataTestShot";

         A     "M_NewShotDataTestShot";
         A     "HT_new_shot_data_valid";
         R     "HT_new_shot_data_valid";
         R     "M_NewShotDataTestShot";
END_REGION

REGION Network 7: Send data to MC
   // Send Data to mouldcarrier 01
         A     "M_WriteShotDataMC_01";
         JCN   MC02;

         CALL  BLKMOV
         ( SRCBLK  := "DB1500_ShotDataToMC".ShotData_MC[0].Data_to_MC,
           RET_VAL := #RetVal,
           DSTBLK  := "DB1500_ShotDataToMC".ShotData_MC[1].Data_to_MC
         );

   // Reset requests / set data valid
         SET;
         R     "M_WriteShotDataMC_01";
         R     "M_NewShotDataToMC_01";
         S     "DB1500_ShotDataToMC".ShotData_MC[1].Data_to_MC.Communication.New_Data;

         JU    del;

   // Send Data to mouldcarrier 02
   MC02: A     "M_WriteShotDataMC_02";
         JCN   MC03;

         CALL  BLKMOV
         ( SRCBLK  := "DB1500_ShotDataToMC".ShotData_MC[0].Data_to_MC,
           RET_VAL := #RetVal,
           DSTBLK  := "DB1500_ShotDataToMC".ShotData_MC[2].Data_to_MC
         );

   // Reset requests / set data valid
         SET;
         R     "M_WriteShotDataMC_02";
         R     "M_NewShotDataToMC_02";
         S     "DB1500_ShotDataToMC".ShotData_MC[2].Data_to_MC.Communication.New_Data;

         JU    del;

   // Send Data to mouldcarrier 03
   MC03: A     "M_WriteShotDataMC_03";
         JCN   MC04;

         CALL  BLKMOV
         ( SRCBLK  := "DB1500_ShotDataToMC".ShotData_MC[0].Data_to_MC,
           RET_VAL := #RetVal,
           DSTBLK  := "DB1500_ShotDataToMC".ShotData_MC[3].Data_to_MC
         );

   // Reset requests / set data valid
         SET;
         R     "M_WriteShotDataMC_03";
         R     "M_NewShotDataToMC_03";
         S     "DB1500_ShotDataToMC".ShotData_MC[3].Data_to_MC.Communication.New_Data;

         JU    del;

   // Send Data to mouldcarrier 04
   MC04: A     "M_WriteShotDataMC_04";
         JCN   MC05;

         CALL  BLKMOV
         ( SRCBLK  := "DB1500_ShotDataToMC".ShotData_MC[0].Data_to_MC,
           RET_VAL := #RetVal,
           DSTBLK  := "DB1500_ShotDataToMC".ShotData_MC[4].Data_to_MC
         );

   // Reset requests / set data valid
         SET;
         R     "M_WriteShotDataMC_04";
         R     "M_NewShotDataToMC_04";
         S     "DB1500_ShotDataToMC".ShotData_MC[4].Data_to_MC.Communication.New_Data;

         JU    del;

   // Send Data to mouldcarrier 05
   MC05: A     "M_WriteShotDataTestShot";
         JC    del;
END_REGION

REGION Network 8: Send act data to MC
         L     "DB608_PV_Metering".Metering[1].Flow.PV_ActV.Value;
         T     "DB1500_ShotDataToMC".ShotData_MC[1].Data_to_MC.Act_value.Comp[1].Flow;
         T     "DB1500_ShotDataToMC".ShotData_MC[2].Data_to_MC.Act_value.Comp[1].Flow;

         L     "DB604_PV_Mixinghead".Mixinghead[1].Pressure_Connection[1].PV_ActV.Value;
         T     "DB1500_ShotDataToMC".ShotData_MC[1].Data_to_MC.Act_value.Comp[1].Pressure_MH;
         T     "DB1500_ShotDataToMC".ShotData_MC[2].Data_to_MC.Act_value.Comp[1].Pressure_MH;

         L     "DB604_PV_Mixinghead".Mixinghead[1].Temperature_Connection[1].PV_ActV.Value;
         T     "DB1500_ShotDataToMC".ShotData_MC[1].Data_to_MC.Act_value.Comp[1].Temperature_MH;
         T     "DB1500_ShotDataToMC".ShotData_MC[2].Data_to_MC.Act_value.Comp[1].Temperature_MH;

         L     "DB608_PV_Metering".Metering[2].Flow.PV_ActV.Value;
         T     "DB1500_ShotDataToMC".ShotData_MC[1].Data_to_MC.Act_value.Comp[2].Flow;
         T     "DB1500_ShotDataToMC".ShotData_MC[2].Data_to_MC.Act_value.Comp[2].Flow;

         L     "DB604_PV_Mixinghead".Mixinghead[1].Pressure_Connection[2].PV_ActV.Value;
         T     "DB1500_ShotDataToMC".ShotData_MC[1].Data_to_MC.Act_value.Comp[2].Pressure_MH;
         T     "DB1500_ShotDataToMC".ShotData_MC[2].Data_to_MC.Act_value.Comp[2].Pressure_MH;

         L     "DB604_PV_Mixinghead".Mixinghead[1].Temperature_Connection[2].PV_ActV.Value;
         T     "DB1500_ShotDataToMC".ShotData_MC[1].Data_to_MC.Act_value.Comp[2].Temperature_MH;
         T     "DB1500_ShotDataToMC".ShotData_MC[2].Data_to_MC.Act_value.Comp[2].Temperature_MH;
END_REGION

REGION Network 9: Delete buffer
   del:  NOP   0;

         L     0;
         T     #nullbyte;

         CALL  FILL
         ( BVAL    := #nullbyte,
           RET_VAL := #RetVal,
           BLK     := "DB1500_ShotDataToMC".ShotData_MC[0].Data_to_MC
         );

         SET;
         R     "HT_new_shot_data_valid";
END_REGION

REGION Network 10: End
   End:  NOP   0;
END_REGION

REGION Network 11: Write data to bus
   // MC1
   //      CALL  DPWR_DAT
   //         LADDR   :="PN-PN-Coupler_PU_MC1~OUT_128_Byte_1"
   //         RECORD  :="DB1500_ShotDataToMC".ShotData_MC[1].Data_to_MC
   //         RET_VAL :=#RetValSFC
   // MC2
   //      CALL  DPWR_DAT
   //         LADDR   :="PN-PN-Coupler_PU_MC2~OUT_128_Byte_1"
   //         RECORD  :="DB1500_ShotDataToMC".ShotData_MC[2].Data_to_MC
   //         RET_VAL :=#RetValSFC
   // MC3
   //    CALL  DPWR_DAT
   //         LADDR   :="PN-PN-Coupler_MC3~OUT_128_Byte_1"
   //         RECORD  :="DB1500_ShotDataToMC".ShotData_MC[3].Data_to_MC
   //         RET_VAL :=#RetValSFC
   //    CALL  DPWR_DAT
   //         LADDR   :="PN-PN-Coupler_MC3~OUT_128_Byte_2"
   //         RECORD  :="DB1500_ShotDataToMC".ShotData_MC[3].Data_to_MC.
   //         RET_VAL :=#RetValSFC
   // MC4
   //    CALL  DPWR_DAT
   //         LADDR   :="PN-PN-Coupler_MC4~OUT_128_Byte_1"
   //         RECORD  :="DB1500_ShotDataToMC".ShotData_MC[4].Data_to_MC
   //         RET_VAL :=#RetValSFC
   //    CALL  DPWR_DAT
   //         LADDR   :="PN-PN-Coupler_MC4~OUT_128_Byte_2"
   //         RECORD  :="DB1500_ShotDataToMC".ShotData_MC[4].Data_to_MC
   //         RET_VAL :=#RetValSFC
END_REGION
END_FUNCTION

FUNCTION "FC1900_IF_Kuka_KRC4" : Void   // FC1900, STL
{ S7_Optimized_Access := 'FALSE' }
VERSION : 0.1
   VAR_INPUT
      IN_PW_INOUT : Int;
      IN_Acknowledge_Fault : Bool;
      IN_Auto_Stop_quitt : Bool;   // Autostopp wurde quittiert
      IN_Motorprotection : Bool;
      IN_MH_Automatic : Bool;   // MK in Automatik
      IN_OM_service : Bool;   // Betriebsart Service
      IN_Cycle_running : Bool;   // Zyklus läuft
      IN_Start_cycle : Bool;   // Start Zyklus
      IN_Release_move_MC : Bool;   // Freigabe für Bewegung in die Form
      IN_Shotrelease : Bool;   // Schussfreigabe
      IN_Shotend : Bool;   // Schussende
      IN_FLT_Group_1 : Bool;   // Störgruppe 1 aktiv
      IN_PGNO_MainPos : Byte;   // Programmnummer für Bewegung in Wartungsposition
      IN_PGNO_Cleaning : Byte;   // Programmnummer für Bewegung zum Reinigen
      IN_Timer_Auto_on : Timer;
      IN_Timer_Fault_quitt : Timer;
      IN_Timer_Auto_On_Off : Timer;
      IN_Timer_Delay_Start : Timer;
      IN_Timer_PGNO_Valid : Timer;
      IN_Timer_Imp_ExtStart : Timer;
      AB_KUKA_PGNO : Byte;
   END_VAR
   VAR_IN_OUT
      IO_Button_MainPos : Bool;   // Schalter Wartungsposition
      IO_Button_Cleaning : Bool;   // Schalter Reinigen
      IO_State_MainPos : Byte;   // Status Wartungsposition
      IO_State_Cleaning : Byte;   // Status Reinigen
      IO_Status : "Kuka_KRC4_Status";
      IO_NewFault : Bool;
      IO_FaultLevel_3 : Bool;
   END_VAR
   VAR_TEMP
      Temp_IO_Status : "Kuka_KRC4_Status";
      Anyzeiger : ANY;
      ERROR_CODE : Int;
      Schleifenzaehler : Int;
      Prog_Nummer : Byte;
   END_VAR
BEGIN

REGION Network 1: Gesicherte Daten einbinden
   //----
         LAR1;
         L;
         LAR2;
   //----
         L     W#16#1002;  // Bytes
         T     W [AR1,P#0.0];
         L     36;  // Anzahl Bytes
         T     W [AR1,P#2.0];
         L     W [AR2,P#0.0];  // Baustein Nr.
         T     W [AR1,P#4.0];
         L     D [AR2,P#2.0];  // Datenanfang
         T     D [AR1,P#6.0];
   //----
         CALL  BLKMOV
         ( SRCBLK  := #Anyzeiger,
           RET_VAL := #ERROR_CODE,
           DSTBLK  := #Temp_IO_Status
         );
   //----
END_REGION

REGION Network 2: Ausgänge von dem Roboter in die Steuerung laden
         L;
         LAR2;
         L     #IN_PW_INOUT;
         SLD   3;
         LAR1;
   //
         L     3;  // Anzahl der Eingangsworte
   Pelp: T     #Schleifenzaehler;
   //
         L     PIW [AR1,P#0.0];  // Eingangsswort
         T     LW [ AR2 , P#24.0 ];  // Eingänge im UDT
   //
         +AR1  P#2.0;
         +AR2  P#2.0;
   //
         L     #Schleifenzaehler;
         LOOP  Pelp;
END_REGION

REGION Network 3: Störungsbehandlung
         A     #IN_Acknowledge_Fault;
         R     #Temp_IO_Status.STG_System;
         R     #Temp_IO_Status.STG_Schnittstelle;
         R     #Temp_IO_Status.STG_Roboter_stoppt;
         R     #Temp_IO_Status.STG_Motoschutz;
   //----
   // Störung KUKA hat gestoppt
         A     #Temp_IO_Status.Input_From_Robot.E_KRC_PRO_ACT;
         FN    #Temp_IO_Status.FHM_PRO_ACT;
         A     #Temp_IO_Status.Input_From_Robot.E_KRC_AUT_EXTERN;
         A     #Temp_IO_Status.Anforderung_Automatik;
         AN    #Temp_IO_Status.STG_Roboter_stoppt;
         S     #Temp_IO_Status.STG_Roboter_stoppt;
         S     #IO_NewFault;

   // Status gestört allgemein
         O     #Temp_IO_Status.STG_Roboter_stoppt;
         AN    #Temp_IO_Status.STG_System;
         S     #Temp_IO_Status.STG_System;
         S     #IO_NewFault;

   // Motorschutz
         AN    #IN_Motorprotection;
         AN    #Temp_IO_Status.STG_Motoschutz;
         S     #Temp_IO_Status.STG_Motoschutz;
         S     #IO_NewFault;

   // Level
         O     #Temp_IO_Status.STG_System;
         O     #Temp_IO_Status.STG_Schnittstelle;
         O     #Temp_IO_Status.STG_Roboter_stoppt;
         O     #Temp_IO_Status.STG_Motoschutz;
         S     #IO_FaultLevel_3;

   // STG quitt an KUKA
         A     #Temp_IO_Status.Input_From_Robot.E_KRC_STOPMES;
   //    U     #Temp_IO_Status.Input_From_Robot.E_KRC_PERI_RDY
         A     #Temp_IO_Status.Input_From_Robot.E_KRC_AUT_EXTERN;
         A     #Temp_IO_Status.Anforderung_Automatik;
         L     s5t#500ms;
         SD    #IN_Timer_Fault_quitt;
         A     #IN_Timer_Fault_quitt;
         =     #Temp_IO_Status.Output_To_Robot.A_SPS_CONF_MESS;
END_REGION

REGION Network 4: Roboter starten und stoppen
   //----
   // Antriebe einschalten
   //----
         A     #Temp_IO_Status.Input_From_Robot.E_KRC_AUT_EXTERN;
         A     #Temp_IO_Status.Input_From_Robot.E_KRC_USER_SAF;
         A     #Temp_IO_Status.Input_From_Robot.E_KRC_ALARM_STOP;
         A     #IN_MH_Automatic;
         AN    #Temp_IO_Status.STG_System;
         AN    #Temp_IO_Status.STG_Schnittstelle;
         AN    #Temp_IO_Status.STG_Roboter_stoppt;
         =     #Temp_IO_Status.Anforderung_Automatik;
   //----
         A     #Temp_IO_Status.Anforderung_Automatik;
         L     S5T#500MS;
         SD    #IN_Timer_Auto_on;
   //----
         A     #Temp_IO_Status.Anforderung_Automatik;
         =     #Temp_IO_Status.Output_To_Robot.A_SPS_DRIVES_OFF;
   //----
         A     #IN_Timer_Auto_on;
         A     #Temp_IO_Status.Anforderung_Automatik;
         AN    #Temp_IO_Status.Input_From_Robot.E_KRC_PERI_RDY;
         =     #Temp_IO_Status.Output_To_Robot.A_SPS_DRIVES_ON;
   //----
   // Bewegungsfreigabe
   //----
         A     #Temp_IO_Status.Anforderung_Automatik;
         O     #Temp_IO_Status.Input_From_Robot.E_KRC_T1;
         O     #Temp_IO_Status.Input_From_Robot.E_KRC_T2;
         =     #Temp_IO_Status.Output_To_Robot.A_SPS_MOVE_ENABLE;
   //----
   // Prozess starten
   //----
         A     #Temp_IO_Status.Anforderung_Automatik;
         A     #Temp_IO_Status.Input_From_Robot.E_KRC_PERI_RDY;
   //   U(
   //      O     #Temp_IO_Status.Input_From_Robot.E_KRC_IN_HOME
   //      O(
   //      U     #Temp_IO_Status.Input_From_Robot.E_KRC_IN_MAINPOS
   //      UN    #IN_Cycle_running
   //      )
   //      )
         AN    #Temp_IO_Status.Input_From_Robot.E_KRC_PRO_ACT;
         AN    #Temp_IO_Status.Input_From_Robot.E_KRC_STOPMES;
         =     #Temp_IO_Status.Output_To_Robot.A_SPS_EXT_START;  // Bis zur Loop Schleife im Cell
END_REGION

REGION Network 5: Roboter Positionen // MainPos, Reinigen
   // Während Zyklus Button ablöschen
         A     #IN_Cycle_running;
         AN    #Temp_IO_Status.Input_From_Robot.E_KRC_IN_HOME;
         R     #IO_Button_MainPos;
         R     #IO_Button_Cleaning;

         A     #Temp_IO_Status.Output_To_Robot.A_SPS_INTERRUPT;
         R     #IO_Button_MainPos;

   // HomePos To MainPos
         A     #IO_Button_MainPos;
   //   FP    #Temp_IO_Status.FHM_MainPosToHomePos
         AN    #IN_Cycle_running;
         A     #Temp_IO_Status.Input_From_Robot.E_KRC_IN_HOME;
         A     #Temp_IO_Status.Anforderung_Automatik;
         JCN   MainPos;
         L     #IN_PGNO_MainPos;
         T     #Temp_IO_Status.A_SPS_PGNO;
   MainPos:NOP   0;

   // MainPos to HomePos
         AN    #IO_Button_MainPos;
         A     #Temp_IO_Status.Input_From_Robot.E_KRC_IN_MAINPOS;
         A     #Temp_IO_Status.Anforderung_Automatik;
         =     #Temp_IO_Status.Output_To_Robot.A_KRC_MOVE_TO_HOMEPOS;
   //-----
   // Cleaning MH
         A     #IO_Button_Cleaning;
   //    FP    #Temp_IO_Status.FHM_Cleaning_MH
         AN    #IN_Cycle_running;
         A     #Temp_IO_Status.Input_From_Robot.E_KRC_IN_HOME;
         A     #Temp_IO_Status.Anforderung_Automatik;
         JCN   Cleaning;
         L     #IN_PGNO_Cleaning;
         T     #Temp_IO_Status.A_SPS_PGNO;
   Cleaning:NOP   0;

         A     #IO_Button_Cleaning;
         AN    #Temp_IO_Status.Input_From_Robot.E_KRC_IN_HOME;
         R     #IO_Button_Cleaning;
   //-----
   // Status MainPos

         L     1;
         A     #IO_Button_MainPos;
         A     #Temp_IO_Status.Input_From_Robot.E_KRC_IN_MAINPOS;
         JC    StateMainPos;

         L     3;
         A     #IO_Button_MainPos;
         AN    #Temp_IO_Status.Input_From_Robot.E_KRC_IN_MAINPOS;
         JC    StateMainPos;

         L     0;
   StateMainPos:T     #IO_State_MainPos;
   //-----
   // Status cleaning

         L     1;
         A     #IO_Button_Cleaning;
         JC    Statecleaning;

         L     0;
   Statecleaning:T     #IO_State_Cleaning;
END_REGION

